(* Logix 5000 project; controller FV vendor 1 type 14 code 217 rev 31.11; software revision 31.00; part 17 of 63 *)
(* tags used below, declared in another part *)
   CWD : CHECKWORD_FLAGS;
   FR_data_file_value_to_move : DINT;
   FR_FV26_AV05 : PlantItem;   // FV26_AV05
   FR_FV27_AV05 : PlantItem;   // FV27_AV05
   FR_FV28_AV05 : PlantItem;   // FV28_AV05
   FR_FV29_AV05 : PlantItem;   // FV29_AV05
   FR_GBM_P01 : PlantItem;   // GBM_P01
   FR_N100 : INT[265];   // FV FILLING
   FR_N110 : INT[265];   // GREEN BEER Green Beer Main
   FR_N120 : INT[265];   // YEAST CROP Yeast Cropping Main
   FR_N13 : INT[265];   // MV_ROUTE Comms to MV Routing PLC
   FR_N130 : INT[265];   // FILTRATE Filtrate Return
   FR_N14 : INT[265];   // MVFV CIP Comms to MVFV CIP Un it PLC
   FR_N140 : INT[265];   // CIP
   FR_N160 : INT[265];   // VESSEL Vessel Working Direc tory
   FR_N255 : INT[265];   // CHECKWORDS
   FR_N26 : INT[265];   // FV26
   FR_N27 : INT[265];   // FV27
   FR_N28 : INT[265];   // FV28
   FR_N29 : INT[265];   // FV29
   FR_N30 : INT[265];   // FV30
   FR_N31 : INT[265];   // FV31
   FR_N99 : INT[265];   // COMMENT Comment Lines
   FR_PANELESTOP : PlantItem;   // PANELESTOP
   FR_PILZ : PlantItem;   // PILZ
   FR_T111 : TIMER[255];   // GREEN BEER
   FR_T144 : TIMER[255];   // CIP
   FR_VB1_AV01 : PlantItem;   // VB1_AV01
   FR_VB1_AV03 : PlantItem;   // VB1_AV03
   FR_VB1_AV06 : PlantItem;   // VB1_AV06
   FR_VB2_AV02 : PlantItem;   // VB2_AV02
   FR_VB3_AV02 : PlantItem;   // VB3_AV02
   FR_YP1_CIPRET : PlantItem;   // YP1_CIPRET
   FR_YP2_CIPRET : PlantItem;   // YP2_CIPRET
   FR_YP3_CIPRET : PlantItem;   // YP3_CIPRET
(* FR_Common, continued *)

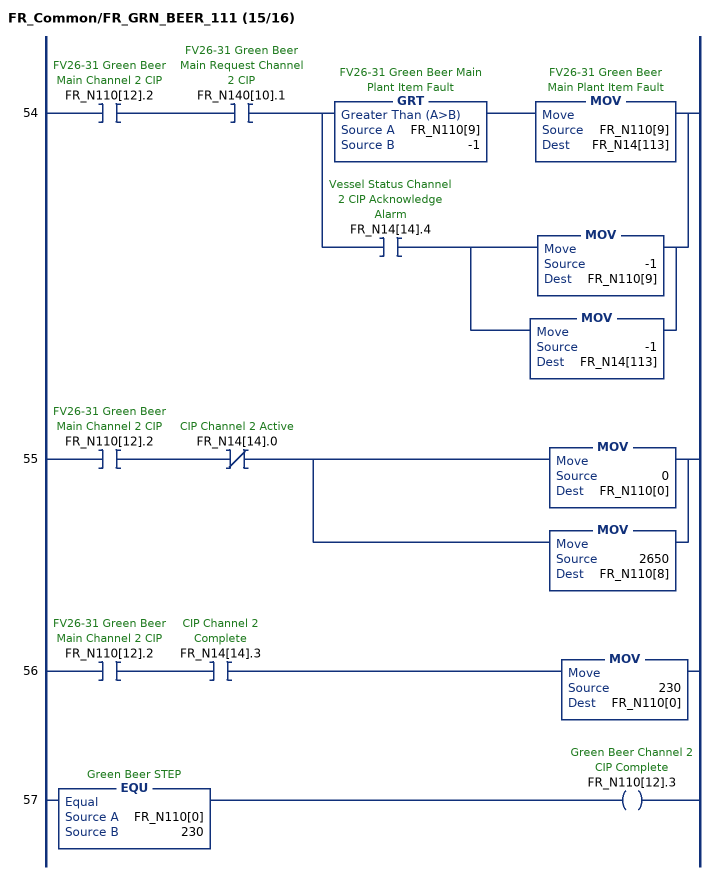
   [picture p273: FR_Common/FR_GRN_BEER_111 rungs 54-57]
   54: XIC(FR_N110[12].2)XIC(FR_N140[10].1)[GRT(FR_N110[9],-1) MOV(FR_N110[9],FR_N14[113]) ,XIC(FR_N14[14].4) [MOV(-1,FR_N110[9]) ,MOV(-1,FR_N14[113]) ] ];
   55: XIC(FR_N110[12].2)XIO(FR_N14[14].0)[MOV(0,FR_N110[0]) ,MOV(2650,FR_N110[8]) ];
   56: XIC(FR_N110[12].2)XIC(FR_N14[14].3)MOV(230,FR_N110[0]);
   57: EQU(FR_N110[0],230)OTE(FR_N110[12].3);
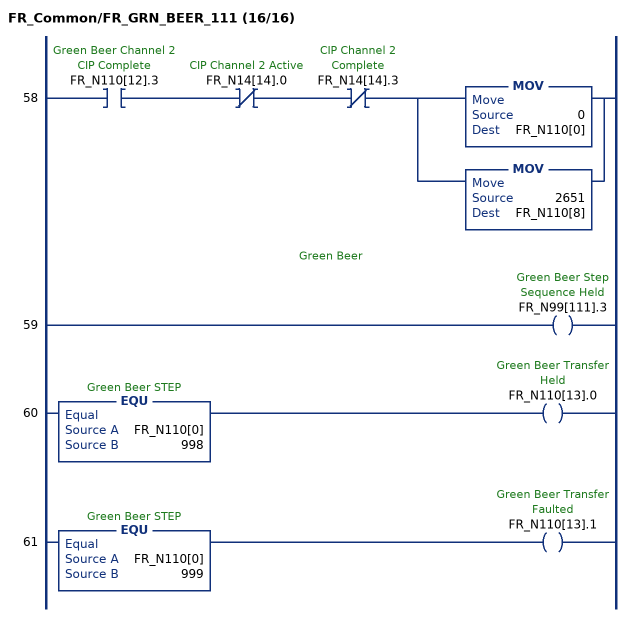
   58: XIC(FR_N110[12].3)XIO(FR_N14[14].0)XIO(FR_N14[14].3)[MOV(0,FR_N110[0]) ,MOV(2651,FR_N110[8]) ];
   // Green Beer
   59: OTE(FR_N99[111].3);
   60: EQU(FR_N110[0],998)OTE(FR_N110[13].0);
   61: EQU(FR_N110[0],999)OTE(FR_N110[13].1);
END_ROUTINE

ROUTINE FR_GRN_BEEROP_112   (* ladder *)
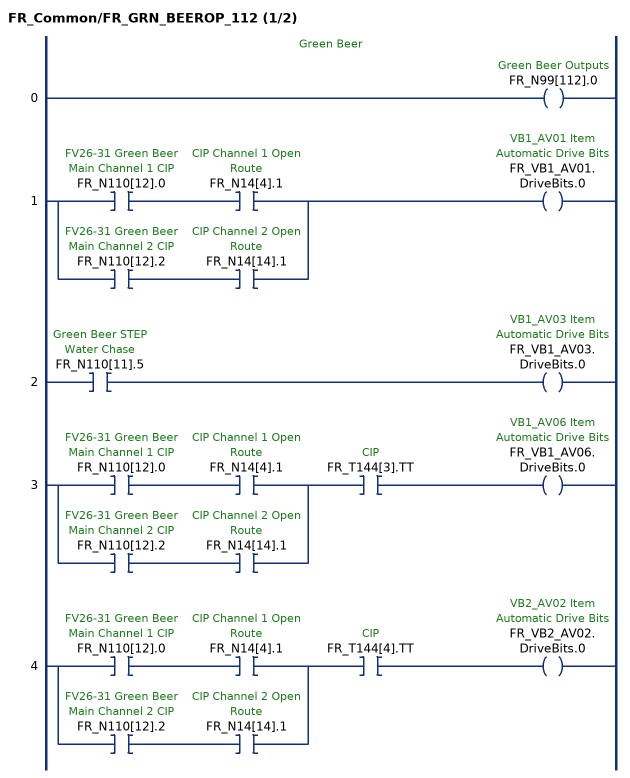
   // Green Beer
   0: OTE(FR_N99[112].0);
   1: [XIC(FR_N110[12].0) XIC(FR_N14[4].1) ,XIC(FR_N110[12].2) XIC(FR_N14[14].1) ]OTE(FR_VB1_AV01.DriveBits.0);
   2: XIC(FR_N110[11].5)OTE(FR_VB1_AV03.DriveBits.0);
   3: [XIC(FR_N110[12].0) XIC(FR_N14[4].1) ,XIC(FR_N110[12].2) XIC(FR_N14[14].1) ]XIC(FR_T144[3].TT)OTE(FR_VB1_AV06.DriveBits.0);
   4: [XIC(FR_N110[12].0) XIC(FR_N14[4].1) ,XIC(FR_N110[12].2) XIC(FR_N14[14].1) ]XIC(FR_T144[4].TT)OTE(FR_VB2_AV02.DriveBits.0);
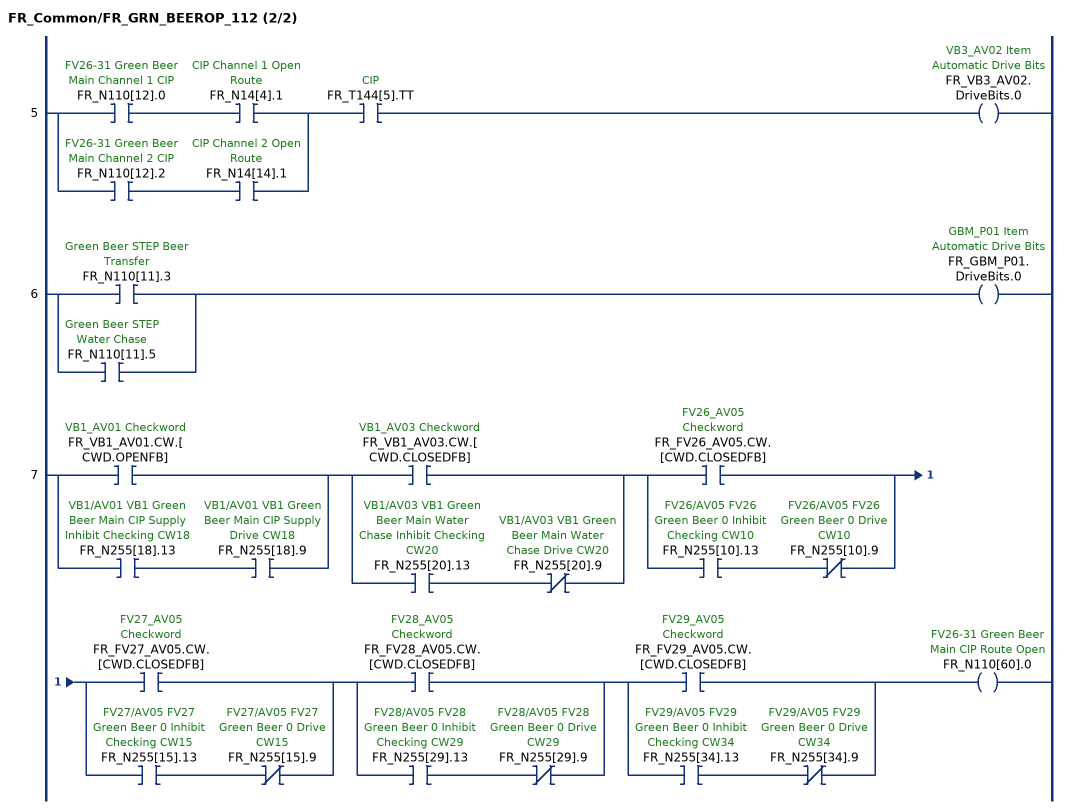
   5: [XIC(FR_N110[12].0) XIC(FR_N14[4].1) ,XIC(FR_N110[12].2) XIC(FR_N14[14].1) ]XIC(FR_T144[5].TT)OTE(FR_VB3_AV02.DriveBits.0);
   6: [XIC(FR_N110[11].3) ,XIC(FR_N110[11].5) ]OTE(FR_GBM_P01.DriveBits.0);
   7: [XIC(FR_VB1_AV01.CW.[CWD.OPENFB]) ,XIC(FR_N255[18].13) XIC(FR_N255[18].9) ][XIC(FR_VB1_AV03.CW.[CWD.CLOSEDFB]) ,XIC(FR_N255[20].13) XIO(FR_N255[20].9) ][XIC(FR_FV26_AV05.CW.[CWD.CLOSEDFB]) ,XIC(FR_N255[10].13) XIO(FR_N255[10].9) ][XIC(FR_FV27_AV05.CW.[CWD.CLOSEDFB]) ,XIC(FR_N255[15].13) XIO(FR_N255[15].9) ][XIC(FR_FV28_AV05.CW.[CWD.CLOSEDFB]) ,XIC(FR_N255[29].13) XIO(FR_N255[29].9) ][XIC(FR_FV29_AV05.CW.[CWD.CLOSEDFB]) ,XIC(FR_N255[34].13) XIO(FR_N255[34].9) ]OTE(FR_N110[60].0);
END_ROUTINE

ROUTINE FR_GRN_BEERST_110   (* ladder *)
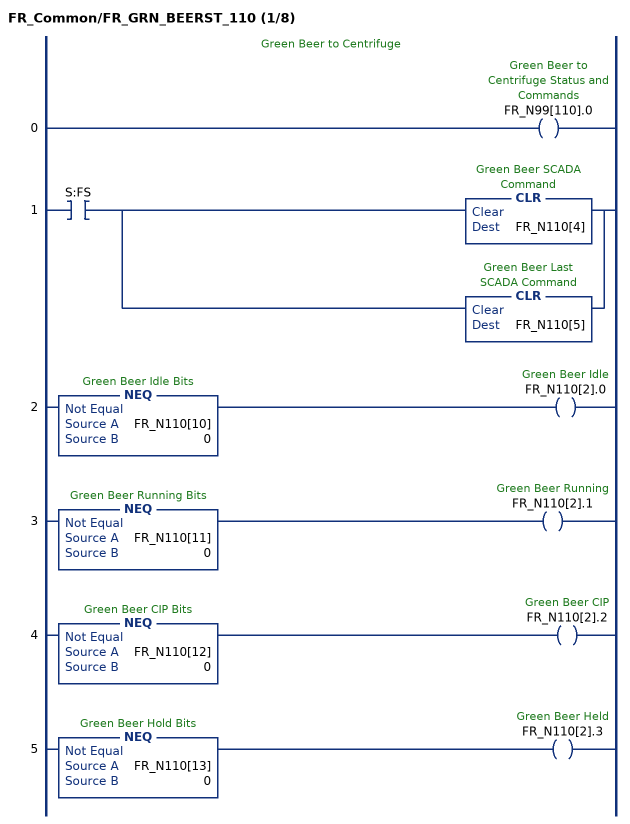
   // Green Beer to Centrifuge
   0: OTE(FR_N99[110].0);
   1: XIC(S:FS)[CLR(FR_N110[4]) ,CLR(FR_N110[5]) ];
   2: NEQ(FR_N110[10],0)OTE(FR_N110[2].0);
   3: NEQ(FR_N110[11],0)OTE(FR_N110[2].1);
   4: NEQ(FR_N110[12],0)OTE(FR_N110[2].2);
   5: NEQ(FR_N110[13],0)OTE(FR_N110[2].3);
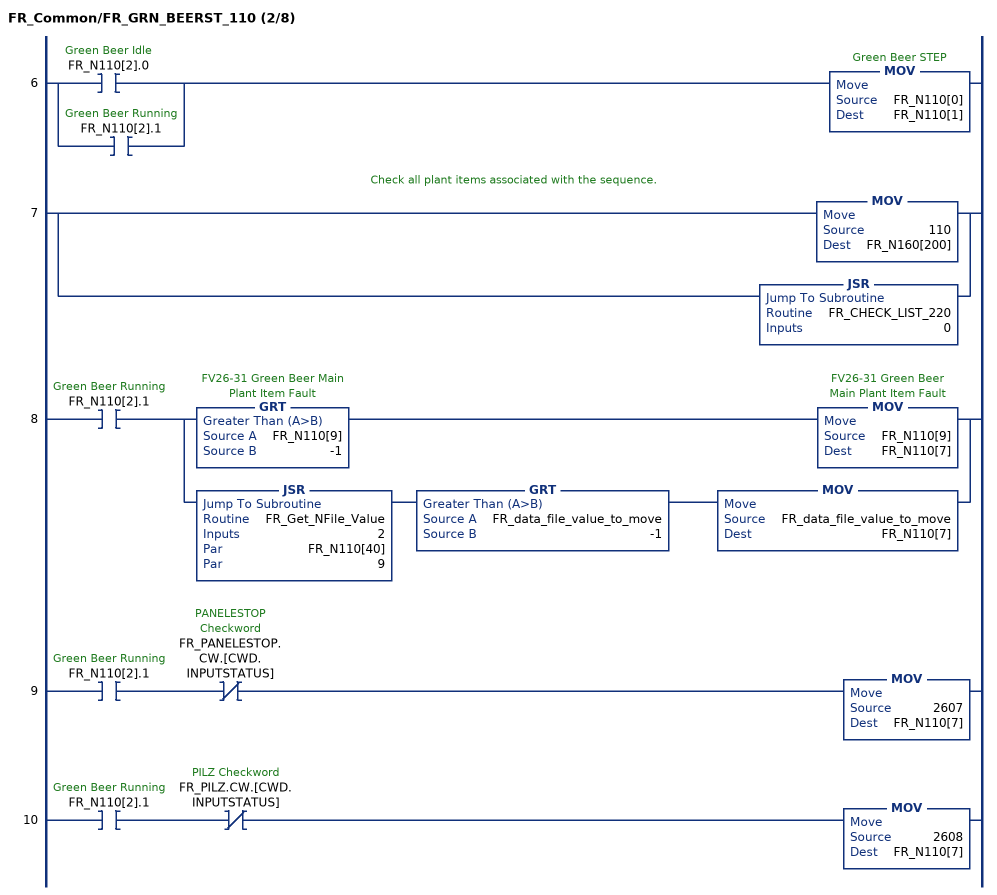
   6: [XIC(FR_N110[2].0) ,XIC(FR_N110[2].1) ]MOV(FR_N110[0],FR_N110[1]);
   // Check all plant items associated with the sequence.
   7: [MOV(110,FR_N160[200]) ,JSR(FR_CHECK_LIST_220,0) ];
   8: XIC(FR_N110[2].1)[GRT(FR_N110[9],-1) MOV(FR_N110[9],FR_N110[7]) ,JSR(FR_Get_NFile_Value,2,FR_N110[40],9) GRT(FR_data_file_value_to_move,-1) MOV(FR_data_file_value_to_move,FR_N110[7]) ];
   9: XIC(FR_N110[2].1)XIO(FR_PANELESTOP.CW.[CWD.INPUTSTATUS])MOV(2607,FR_N110[7]);
   10: XIC(FR_N110[2].1)XIO(FR_PILZ.CW.[CWD.INPUTSTATUS])MOV(2608,FR_N110[7]);
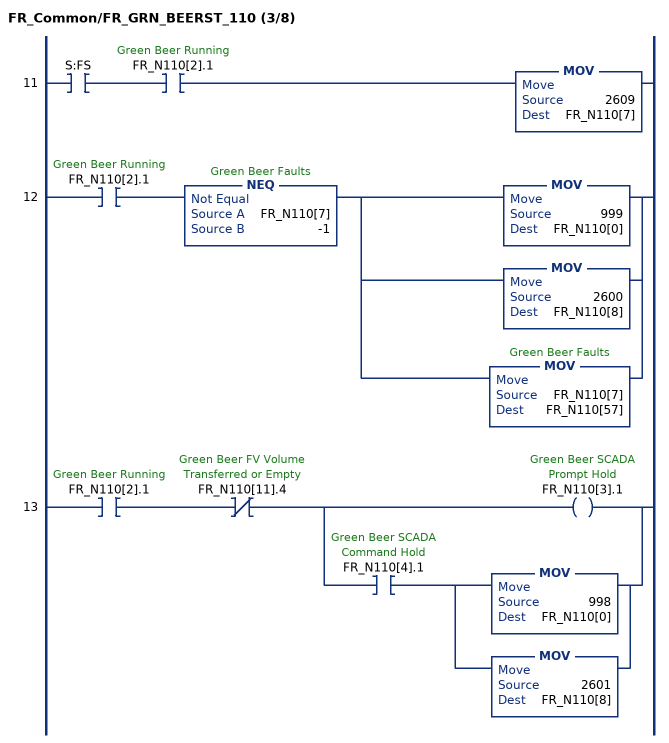
   11: XIC(S:FS)XIC(FR_N110[2].1)MOV(2609,FR_N110[7]);
   12: XIC(FR_N110[2].1)NEQ(FR_N110[7],-1)[MOV(999,FR_N110[0]) ,MOV(2600,FR_N110[8]) ,MOV(FR_N110[7],FR_N110[57]) ];
   13: XIC(FR_N110[2].1)XIO(FR_N110[11].4)[OTE(FR_N110[3].1) ,XIC(FR_N110[4].1) [MOV(998,FR_N110[0]) ,MOV(2601,FR_N110[8]) ] ];
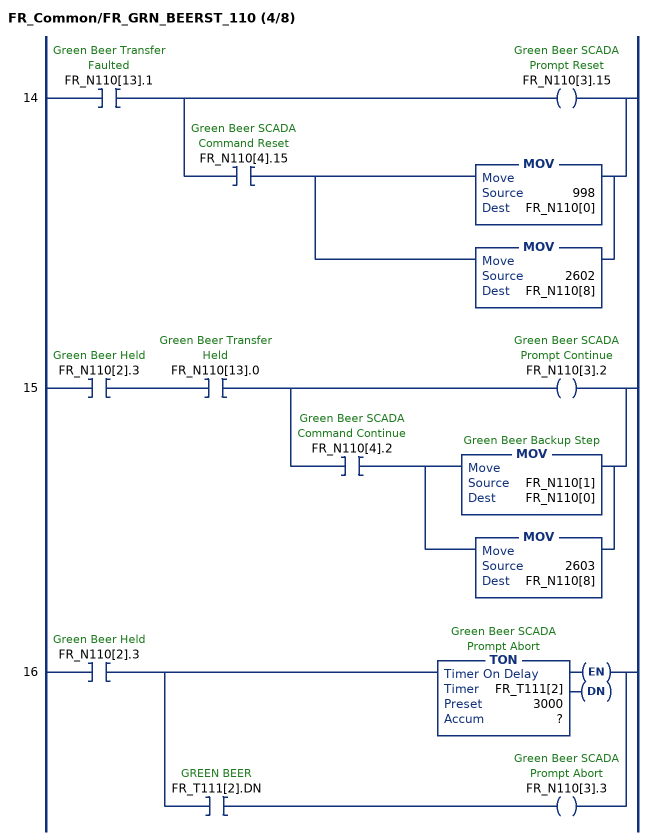
   14: XIC(FR_N110[13].1)[OTE(FR_N110[3].15) ,XIC(FR_N110[4].15) [MOV(998,FR_N110[0]) ,MOV(2602,FR_N110[8]) ] ];
   15: XIC(FR_N110[2].3)XIC(FR_N110[13].0)[OTE(FR_N110[3].2) ,XIC(FR_N110[4].2) [MOV(FR_N110[1],FR_N110[0]) ,MOV(2603,FR_N110[8]) ] ];
   16: XIC(FR_N110[2].3)[TON(FR_T111[2],?,?) ,XIC(FR_T111[2].DN) OTE(FR_N110[3].3) ];
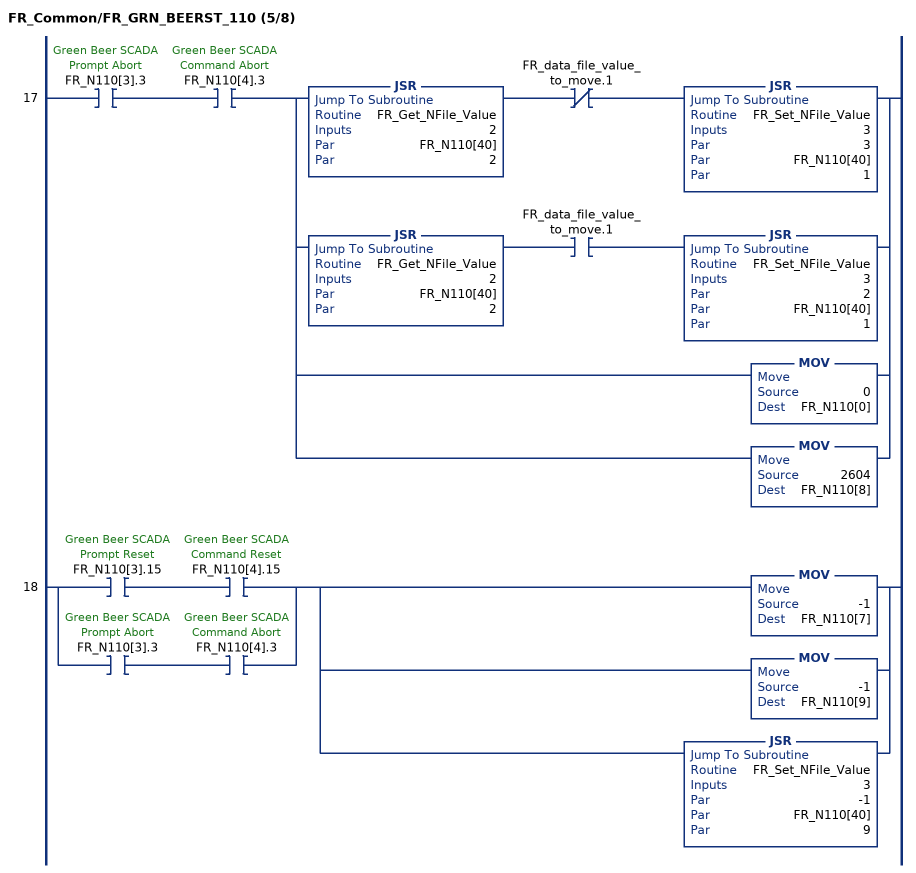
   17: XIC(FR_N110[3].3)XIC(FR_N110[4].3)[JSR(FR_Get_NFile_Value,2,FR_N110[40],2) XIO(FR_data_file_value_to_move.1) JSR(FR_Set_NFile_Value,3,3,FR_N110[40],1) ,JSR(FR_Get_NFile_Value,2,FR_N110[40],2) XIC(FR_data_file_value_to_move.1) JSR(FR_Set_NFile_Value,3,2,FR_N110[40],1) ,MOV(0,FR_N110[0]) ,MOV(2604,FR_N110[8]) ];
   18: [XIC(FR_N110[3].15) XIC(FR_N110[4].15) ,XIC(FR_N110[3].3) XIC(FR_N110[4].3) ][MOV(-1,FR_N110[7]) ,MOV(-1,FR_N110[9]) ,JSR(FR_Set_NFile_Value,3,-1,FR_N110[40],9) ];
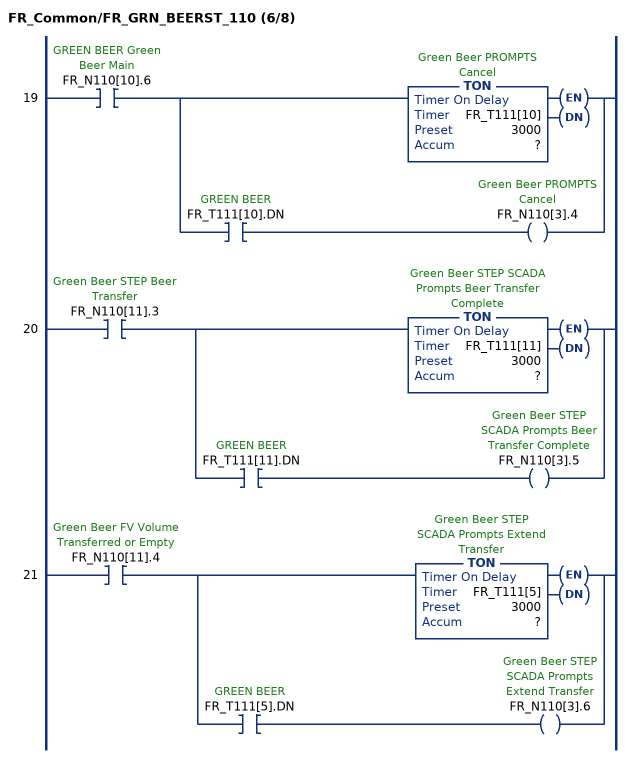
   19: XIC(FR_N110[10].6)[TON(FR_T111[10],?,?) ,XIC(FR_T111[10].DN) OTE(FR_N110[3].4) ];
   20: XIC(FR_N110[11].3)[TON(FR_T111[11],?,?) ,XIC(FR_T111[11].DN) OTE(FR_N110[3].5) ];
   21: XIC(FR_N110[11].4)[TON(FR_T111[5],?,?) ,XIC(FR_T111[5].DN) OTE(FR_N110[3].6) ];
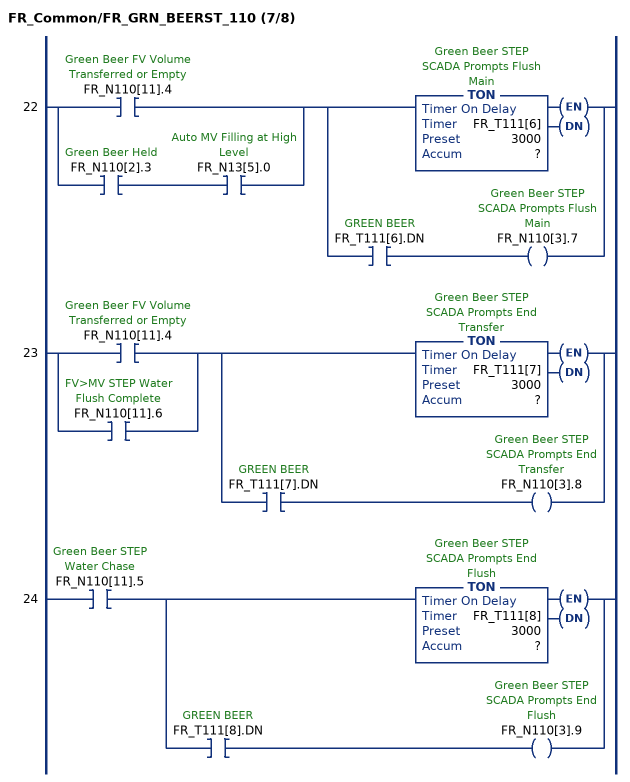
   22: [XIC(FR_N110[11].4) ,XIC(FR_N110[2].3) XIC(FR_N13[5].0) ][TON(FR_T111[6],?,?) ,XIC(FR_T111[6].DN) OTE(FR_N110[3].7) ];
   23: [XIC(FR_N110[11].4) ,XIC(FR_N110[11].6) ][TON(FR_T111[7],?,?) ,XIC(FR_T111[7].DN) OTE(FR_N110[3].8) ];
   24: XIC(FR_N110[11].5)[TON(FR_T111[8],?,?) ,XIC(FR_T111[8].DN) OTE(FR_N110[3].9) ];
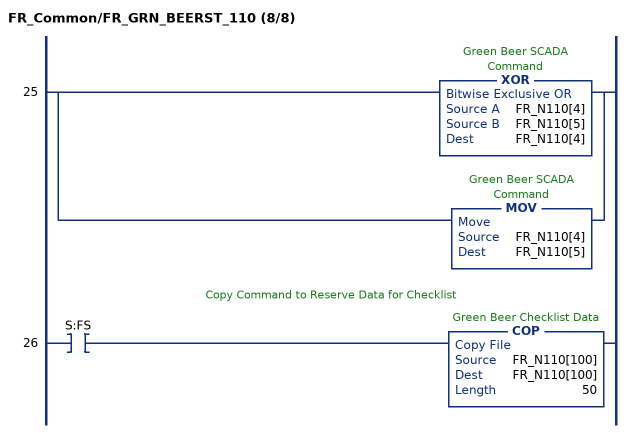
   25: [XOR(FR_N110[4],FR_N110[5],FR_N110[4]) ,MOV(FR_N110[4],FR_N110[5]) ];
   // Copy Command to Reserve Data for Checklist
   26: XIC(S:FS)COP(FR_N110[100],FR_N110[100],50);
END_ROUTINE

ROUTINE FR_INITIALISE_5   (* ladder *)
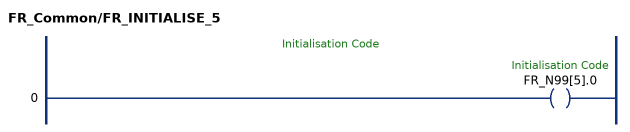
   // Initialisation Code
   0: OTE(FR_N99[5].0);
END_ROUTINE

ROUTINE FR_MVFV_CIP_140   (* ladder *)
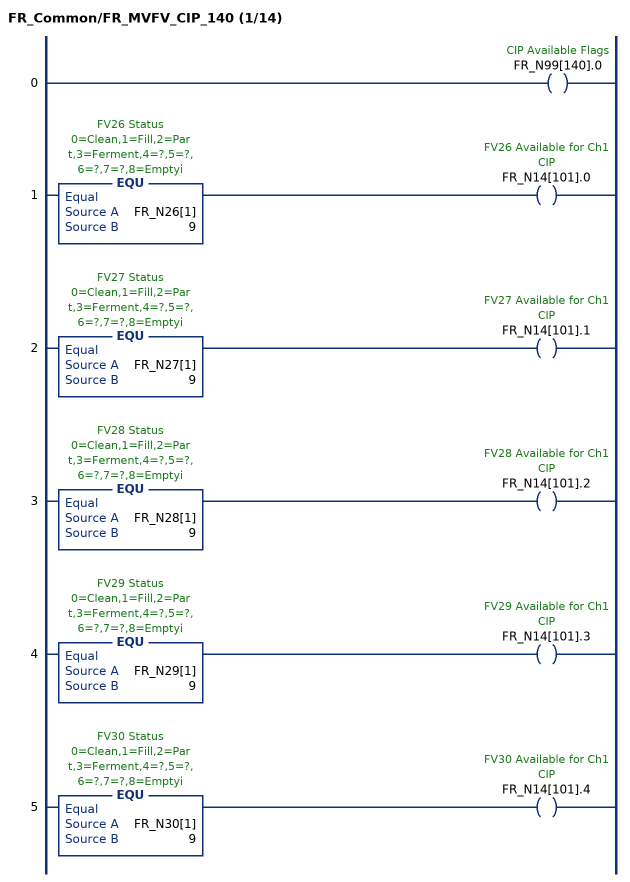
   0: OTE(FR_N99[140].0);
   1: EQU(FR_N26[1],9)OTE(FR_N14[101].0);
   2: EQU(FR_N27[1],9)OTE(FR_N14[101].1);
   3: EQU(FR_N28[1],9)OTE(FR_N14[101].2);
   4: EQU(FR_N29[1],9)OTE(FR_N14[101].3);
   5: EQU(FR_N30[1],9)OTE(FR_N14[101].4);
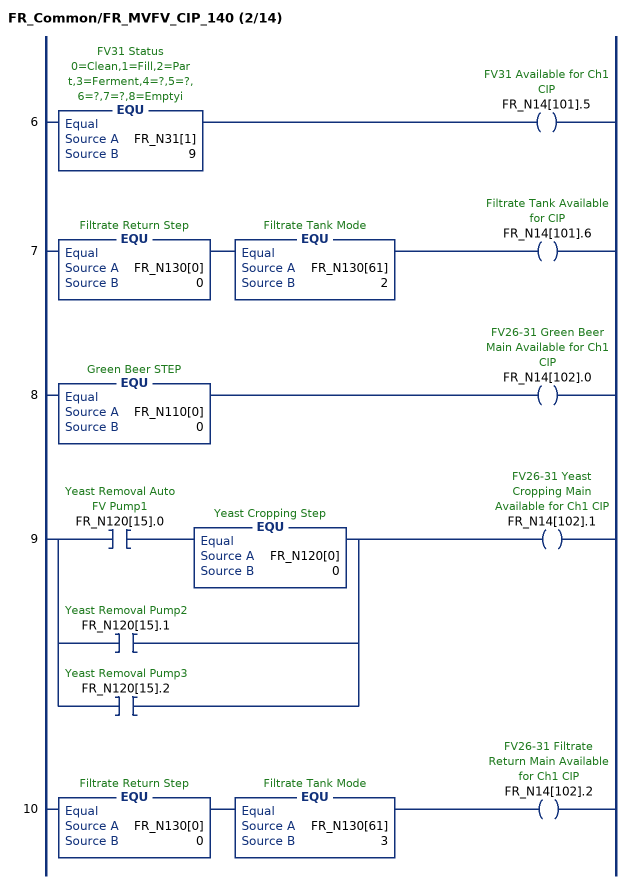
   6: EQU(FR_N31[1],9)OTE(FR_N14[101].5);
   7: EQU(FR_N130[0],0)EQU(FR_N130[61],2)OTE(FR_N14[101].6);
   8: EQU(FR_N110[0],0)OTE(FR_N14[102].0);
   9: [XIC(FR_N120[15].0) EQU(FR_N120[0],0) ,XIC(FR_N120[15].1) ,XIC(FR_N120[15].2) ]OTE(FR_N14[102].1);
   10: EQU(FR_N130[0],0)EQU(FR_N130[61],3)OTE(FR_N14[102].2);
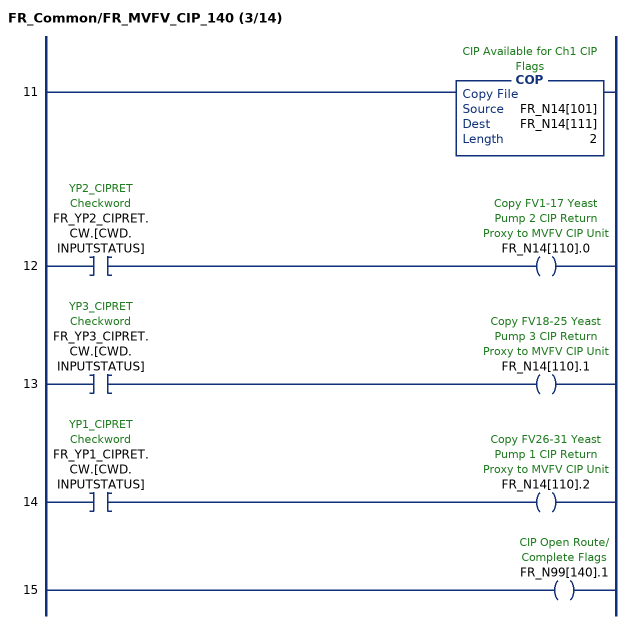
   11: COP(FR_N14[101],FR_N14[111],2);
   12: XIC(FR_YP2_CIPRET.CW.[CWD.INPUTSTATUS])OTE(FR_N14[110].0);
   13: XIC(FR_YP3_CIPRET.CW.[CWD.INPUTSTATUS])OTE(FR_N14[110].1);
   14: XIC(FR_YP1_CIPRET.CW.[CWD.INPUTSTATUS])OTE(FR_N14[110].2);
   15: OTE(FR_N99[140].1);
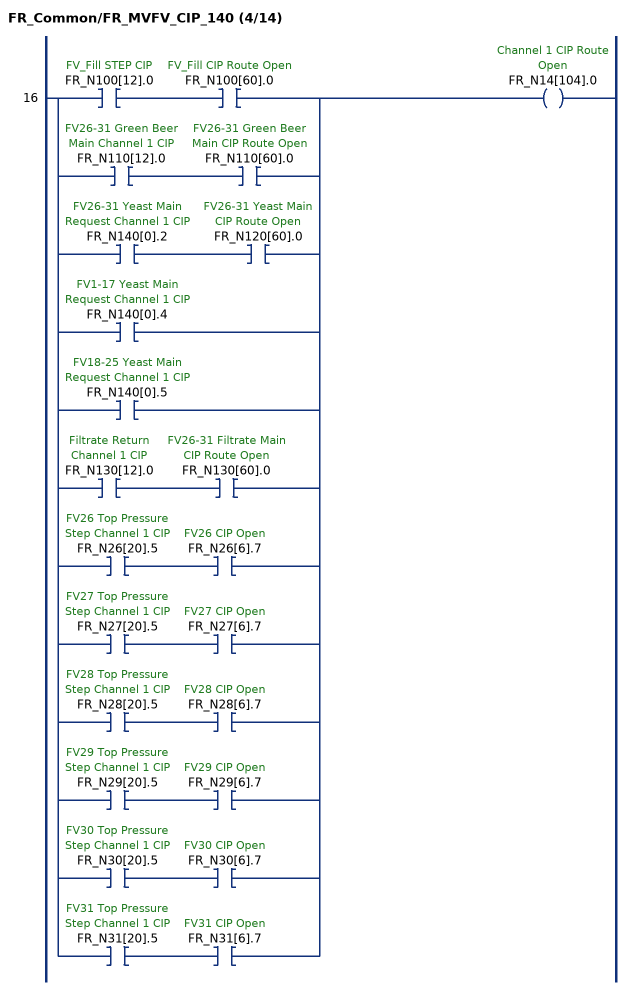
   16: [XIC(FR_N100[12].0) XIC(FR_N100[60].0) ,XIC(FR_N110[12].0) XIC(FR_N110[60].0) ,XIC(FR_N140[0].2) XIC(FR_N120[60].0) ,XIC(FR_N140[0].4) ,XIC(FR_N140[0].5) ,XIC(FR_N130[12].0) XIC(FR_N130[60].0) ,XIC(FR_N26[20].5) XIC(FR_N26[6].7) ,XIC(FR_N27[20].5) XIC(FR_N27[6].7) ,XIC(FR_N28[20].5) XIC(FR_N28[6].7) ,XIC(FR_N29[20].5) XIC(FR_N29[6].7) ,XIC(FR_N30[20].5) XIC(FR_N30[6].7) ,XIC(FR_N31[20].5) XIC(FR_N31[6].7) ]OTE(FR_N14[104].0);
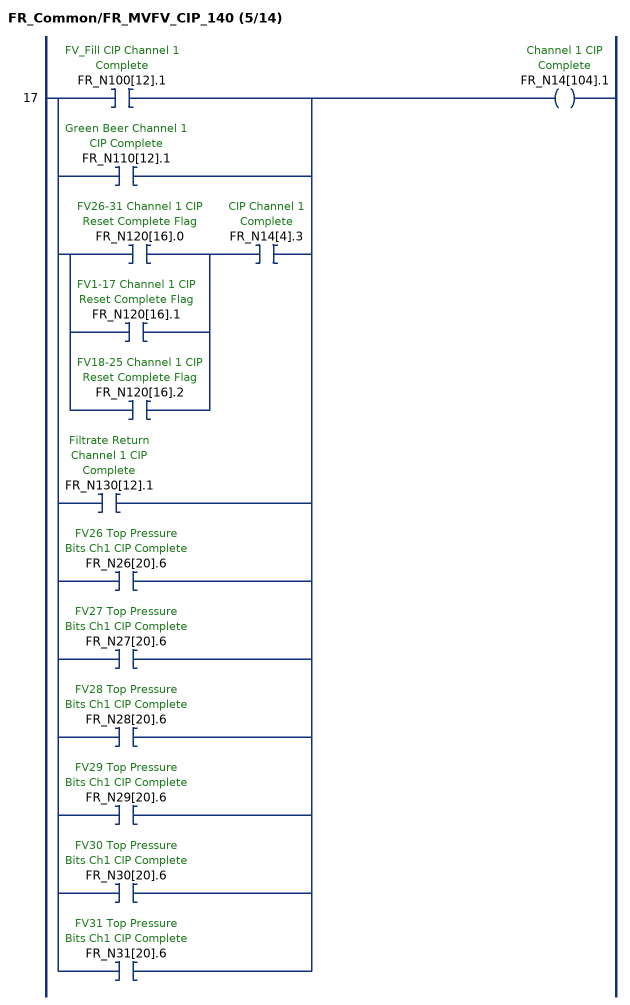
   17: [XIC(FR_N100[12].1) ,XIC(FR_N110[12].1) ,[XIC(FR_N120[16].0) ,XIC(FR_N120[16].1) ,XIC(FR_N120[16].2) ] XIC(FR_N14[4].3) ,XIC(FR_N130[12].1) ,XIC(FR_N26[20].6) ,XIC(FR_N27[20].6) ,XIC(FR_N28[20].6) ,XIC(FR_N29[20].6) ,XIC(FR_N30[20].6) ,XIC(FR_N31[20].6) ]OTE(FR_N14[104].1);
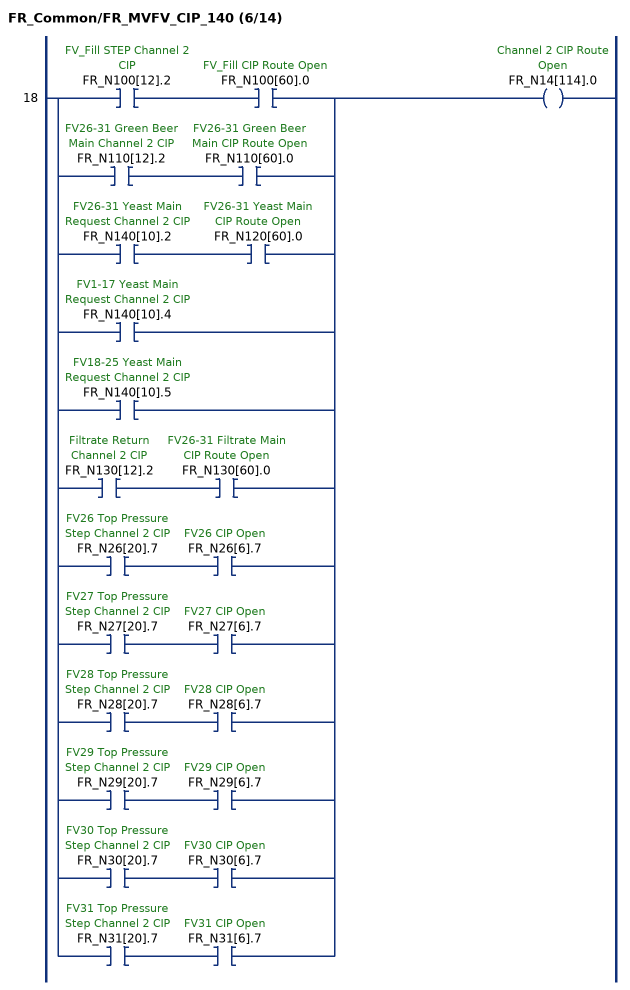
   18: [XIC(FR_N100[12].2) XIC(FR_N100[60].0) ,XIC(FR_N110[12].2) XIC(FR_N110[60].0) ,XIC(FR_N140[10].2) XIC(FR_N120[60].0) ,XIC(FR_N140[10].4) ,XIC(FR_N140[10].5) ,XIC(FR_N130[12].2) XIC(FR_N130[60].0) ,XIC(FR_N26[20].7) XIC(FR_N26[6].7) ,XIC(FR_N27[20].7) XIC(FR_N27[6].7) ,XIC(FR_N28[20].7) XIC(FR_N28[6].7) ,XIC(FR_N29[20].7) XIC(FR_N29[6].7) ,XIC(FR_N30[20].7) XIC(FR_N30[6].7) ,XIC(FR_N31[20].7) XIC(FR_N31[6].7) ]OTE(FR_N14[114].0);
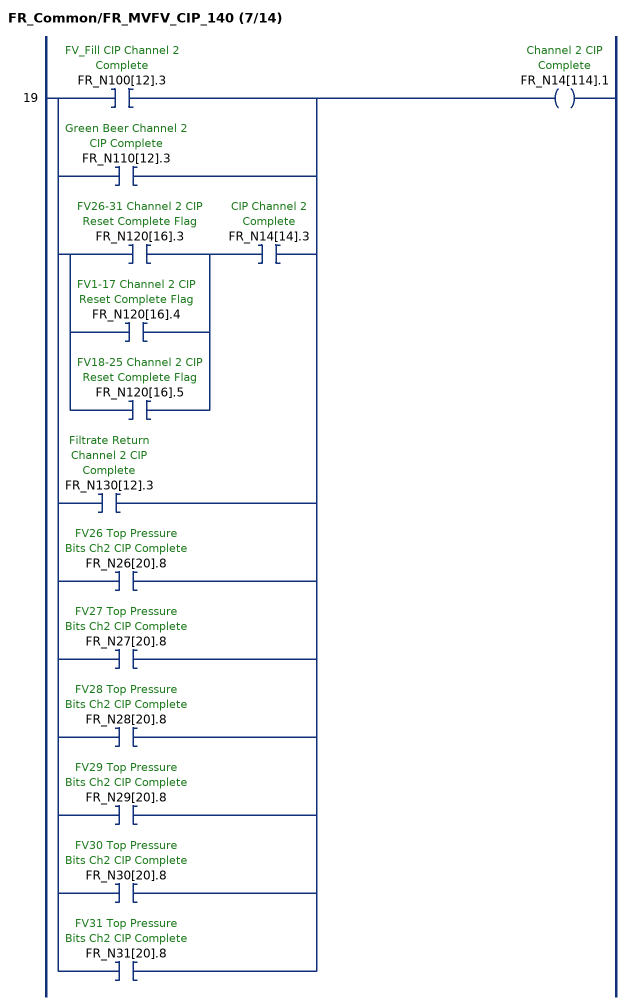
   19: [XIC(FR_N100[12].3) ,XIC(FR_N110[12].3) ,[XIC(FR_N120[16].3) ,XIC(FR_N120[16].4) ,XIC(FR_N120[16].5) ] XIC(FR_N14[14].3) ,XIC(FR_N130[12].3) ,XIC(FR_N26[20].8) ,XIC(FR_N27[20].8) ,XIC(FR_N28[20].8) ,XIC(FR_N29[20].8) ,XIC(FR_N30[20].8) ,XIC(FR_N31[20].8) ]OTE(FR_N14[114].1);
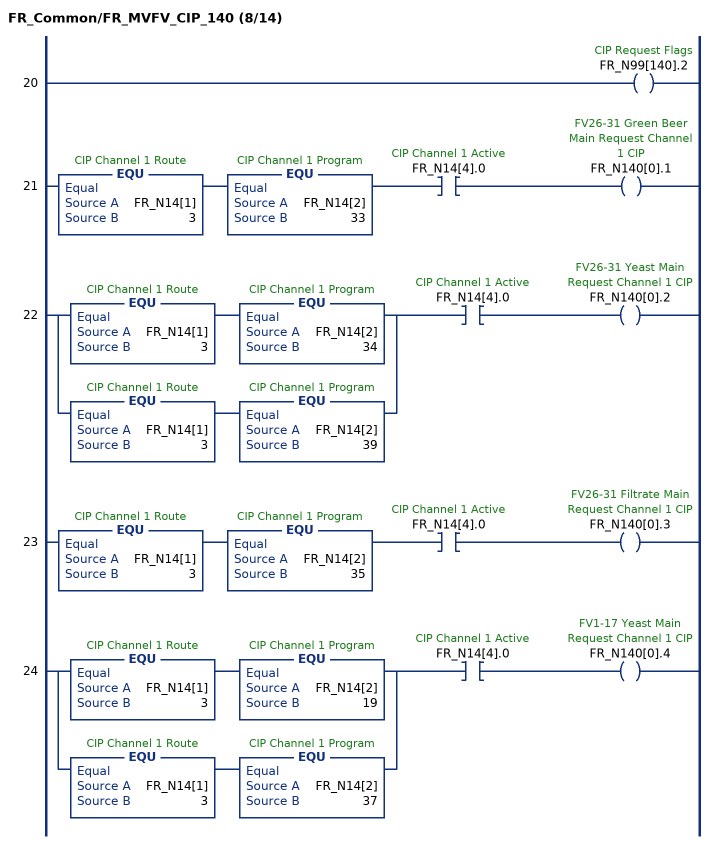
   20: OTE(FR_N99[140].2);
   21: EQU(FR_N14[1],3)EQU(FR_N14[2],33)XIC(FR_N14[4].0)OTE(FR_N140[0].1);
   22: [EQU(FR_N14[1],3) EQU(FR_N14[2],34) ,EQU(FR_N14[1],3) EQU(FR_N14[2],39) ]XIC(FR_N14[4].0)OTE(FR_N140[0].2);
   23: EQU(FR_N14[1],3)EQU(FR_N14[2],35)XIC(FR_N14[4].0)OTE(FR_N140[0].3);
   24: [EQU(FR_N14[1],3) EQU(FR_N14[2],19) ,EQU(FR_N14[1],3) EQU(FR_N14[2],37) ]XIC(FR_N14[4].0)OTE(FR_N140[0].4);
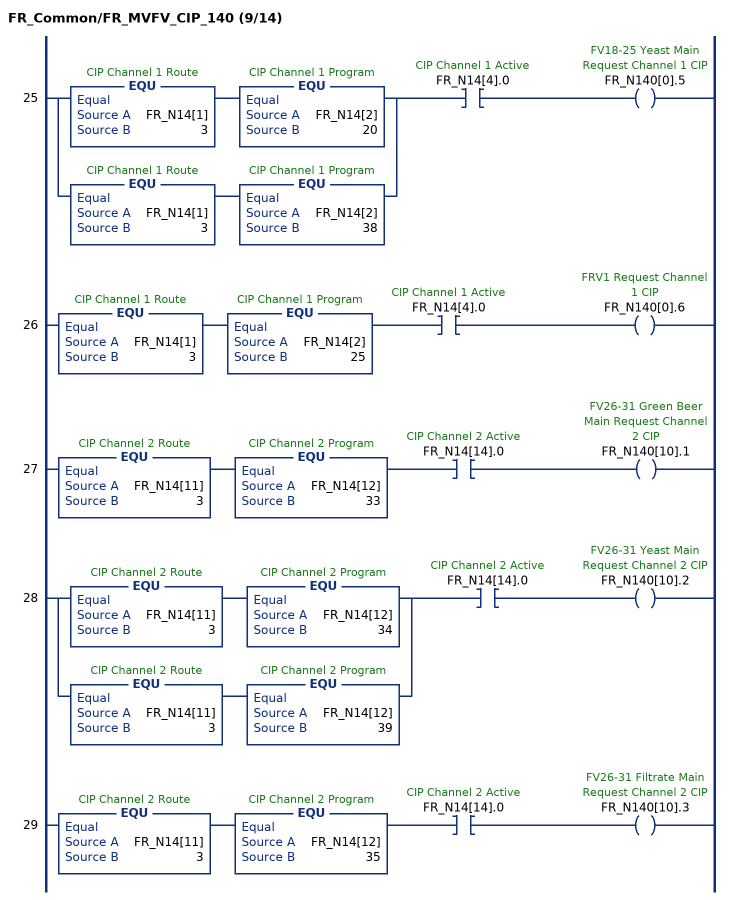
   25: [EQU(FR_N14[1],3) EQU(FR_N14[2],20) ,EQU(FR_N14[1],3) EQU(FR_N14[2],38) ]XIC(FR_N14[4].0)OTE(FR_N140[0].5);
   26: EQU(FR_N14[1],3)EQU(FR_N14[2],25)XIC(FR_N14[4].0)OTE(FR_N140[0].6);
   27: EQU(FR_N14[11],3)EQU(FR_N14[12],33)XIC(FR_N14[14].0)OTE(FR_N140[10].1);
   28: [EQU(FR_N14[11],3) EQU(FR_N14[12],34) ,EQU(FR_N14[11],3) EQU(FR_N14[12],39) ]XIC(FR_N14[14].0)OTE(FR_N140[10].2);
   29: EQU(FR_N14[11],3)EQU(FR_N14[12],35)XIC(FR_N14[14].0)OTE(FR_N140[10].3);
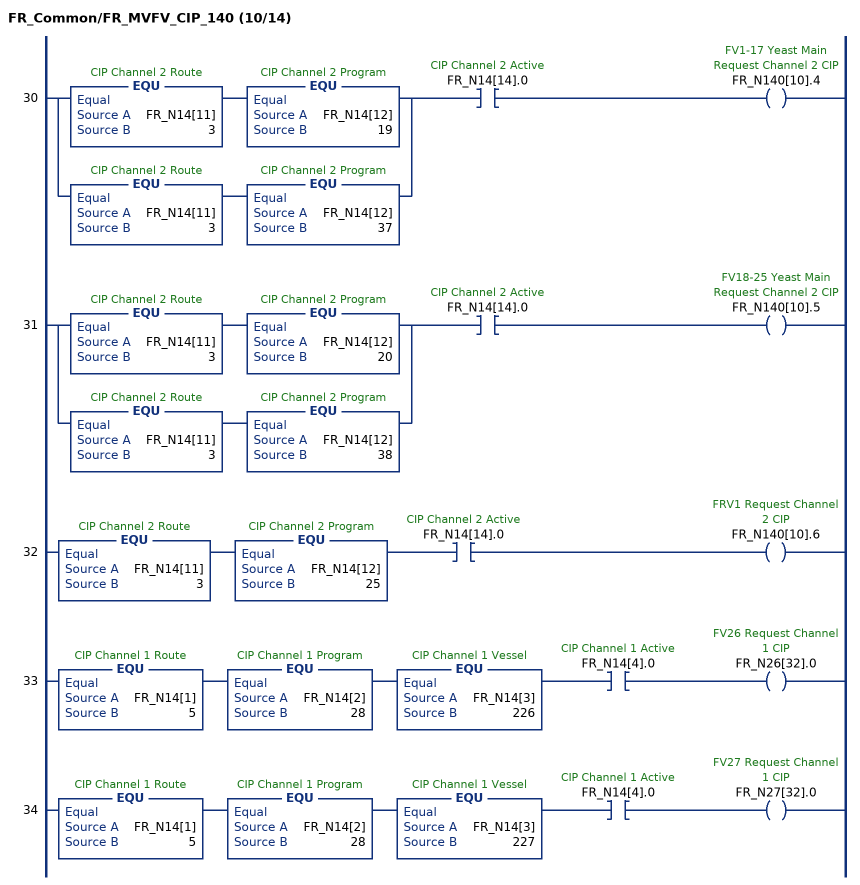
   30: [EQU(FR_N14[11],3) EQU(FR_N14[12],19) ,EQU(FR_N14[11],3) EQU(FR_N14[12],37) ]XIC(FR_N14[14].0)OTE(FR_N140[10].4);
   31: [EQU(FR_N14[11],3) EQU(FR_N14[12],20) ,EQU(FR_N14[11],3) EQU(FR_N14[12],38) ]XIC(FR_N14[14].0)OTE(FR_N140[10].5);
   32: EQU(FR_N14[11],3)EQU(FR_N14[12],25)XIC(FR_N14[14].0)OTE(FR_N140[10].6);
   33: EQU(FR_N14[1],5)EQU(FR_N14[2],28)EQU(FR_N14[3],226)XIC(FR_N14[4].0)OTE(FR_N26[32].0);
   34: EQU(FR_N14[1],5)EQU(FR_N14[2],28)EQU(FR_N14[3],227)XIC(FR_N14[4].0)OTE(FR_N27[32].0);
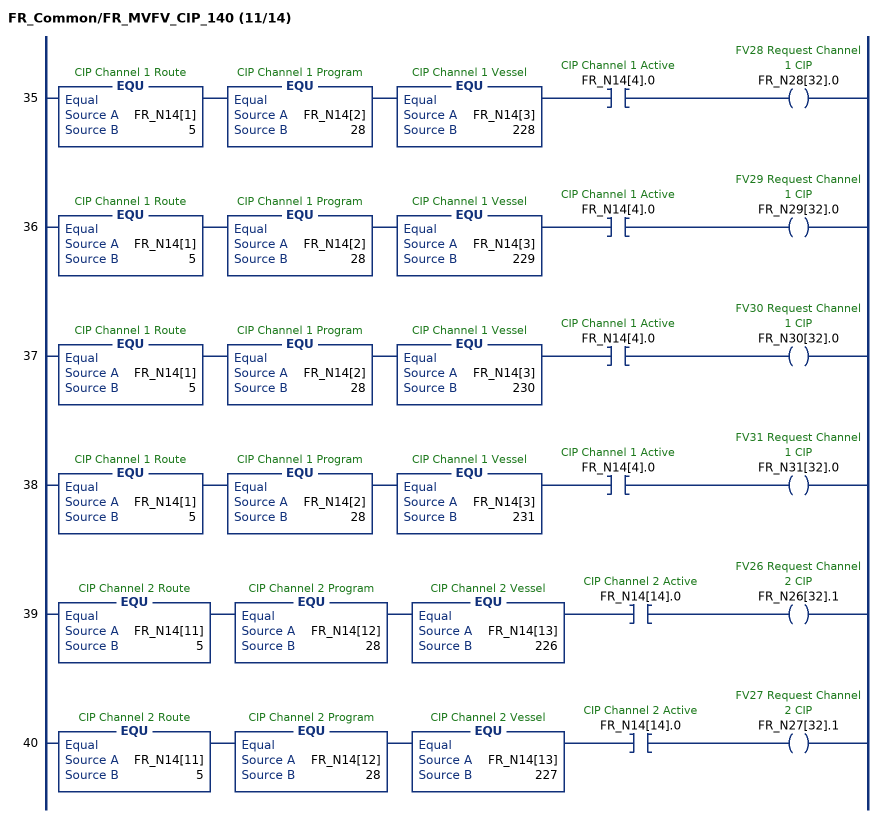
   35: EQU(FR_N14[1],5)EQU(FR_N14[2],28)EQU(FR_N14[3],228)XIC(FR_N14[4].0)OTE(FR_N28[32].0);
   36: EQU(FR_N14[1],5)EQU(FR_N14[2],28)EQU(FR_N14[3],229)XIC(FR_N14[4].0)OTE(FR_N29[32].0);
   37: EQU(FR_N14[1],5)EQU(FR_N14[2],28)EQU(FR_N14[3],230)XIC(FR_N14[4].0)OTE(FR_N30[32].0);
   38: EQU(FR_N14[1],5)EQU(FR_N14[2],28)EQU(FR_N14[3],231)XIC(FR_N14[4].0)OTE(FR_N31[32].0);
   39: EQU(FR_N14[11],5)EQU(FR_N14[12],28)EQU(FR_N14[13],226)XIC(FR_N14[14].0)OTE(FR_N26[32].1);
   40: EQU(FR_N14[11],5)EQU(FR_N14[12],28)EQU(FR_N14[13],227)XIC(FR_N14[14].0)OTE(FR_N27[32].1);
